// TIA Portal project "Symulacja parkingu" (V18)

(* hardware
DEVICE "S7-1200 station_1"  S7-1200 Station
   slot 0: "Rack_0"  S7-1200 Rack  Rack  V1.0
   slot 1: "PLC_1"  CPU 1214C AC/DC/Rly  6ES7 214-1BG40-0XB0  V4.6
DEVICE "HMI_1"  KTP700 Basic PN
   slot 0: "HMI_1"  KTP700 Basic PN  6AV2 123-2GB03-0AX0  17.0.0.0
   slot 1: "HMI_RT_1"  KTP700 Basic PN  6AV2 123-2GB03-0AX0  17.0.0.0
   slot 5: "HMI_1.IE_CP_1"  PROFINET Interface  17.0.0.0
      slot 1: "PROFINET Interface_1"  PROFINET Interface
         slot 1: "Port_1"  Port
*)

// ===== PLC "PLC_1"  CPU 1214C AC/DC/Rly =====

VAR_GLOBAL   // PLC tag table "Default tag table"
   "S1" AT %M0.0 : Bool;   // wjazd
   "S2" AT %M0.1 : Bool;   // wyjazd
   "S3" AT %M0.2 : Bool;   // reset
   "L1" AT %Q0.1 : Bool;   // zielone
   "L2" AT %Q0.2 : Bool;   // czerwone
   "Licznik" AT %MW10 : Word;
   "PV_Wartość_do_ustawienia" AT %MW12 : Word;
   "set wartości do ustawienia" AT %M0.3 : Bool;
   "zmienna do p_triga" AT %M0.4 : Bool;
   "S0" AT %M0.5 : Bool;   // przycisk do całkowitego wyłączenia
   "zmienna pomocnicza do przycisku od wyłączenia" AT %M0.6 : Bool;
   "całkowite wyłączenie" AT %M0.7 : Bool;
   "otwieranie szlabanu wjazd" AT %M1.0 : Bool;
   "otwieranie szlabanu wyjazd" AT %M1.1 : Bool;
   "w trakcie wyjazdu" AT %M1.2 : Bool;
   "w trakcie wjazdu" AT %M1.3 : Bool;
   "L3" AT %M1.4 : Bool;   // pomarańczowy
   "szlaban pozycja wjazd" AT %MW30 : Word;
   "szlaban podnoszenie stan wjazd" AT %M2.0 : Bool;
   "reset timera wjazd podnoszenie" AT %M2.1 : Bool;
   "szlaban opuszczania stan wjazd" AT %M2.2 : Bool;
   "reset timera wjazd opuszczanie" AT %M2.3 : Bool;
   "zmienna pomocnicza do otwierania szlabanu" AT %M2.4 : Bool;
   "szlaban pozycja wyjazd" AT %MW16 : Word;
   "szlaban podnoszenie stan wyjazd" AT %M3.0 : Bool;
   "reset timera wyjazd podnoszenie" AT %M3.1 : Bool;
   "szlaban opuszczania stan wyjazd" AT %M3.2 : Bool;
   "reset timera wyjaazd opuszcanie" AT %M3.3 : Bool;
   "zmienna pomocnicza do otwierania szlabanu 2" AT %M3.4 : Bool;
END_VAR

// folder: System blocks/Program resources

DATA_BLOCK "DB1"   // DB1
{ S7_Optimized_Access := 'TRUE' }
AUTHOR : Simatic
FAMILY : IEC
NAME : CNTR
VERSION : 1.0
// stored: InstanceOfName IEC_COUNTER
"IEC_COUNTER"
BEGIN
END_DATA_BLOCK

DATA_BLOCK "IEC_Timer_0_DB"   // DB2
{ S7_Optimized_Access := 'TRUE' }
AUTHOR : Simatic
FAMILY : IEC
NAME : IEC_TMR
VERSION : 1.0
// stored: InstanceOfName IEC_TIMER
"IEC_TIMER"
BEGIN
END_DATA_BLOCK

DATA_BLOCK "IEC_Timer_0_DB_1"   // DB3
{ S7_Optimized_Access := 'TRUE' }
AUTHOR : Simatic
FAMILY : IEC
NAME : IEC_TMR
VERSION : 1.0
// stored: InstanceOfName IEC_TIMER
"IEC_TIMER"
BEGIN
END_DATA_BLOCK

DATA_BLOCK "IEC_Timer_0_DB_2"   // DB4
{ S7_Optimized_Access := 'TRUE' }
AUTHOR : Simatic
FAMILY : IEC
NAME : IEC_TMR
VERSION : 1.0
// stored: InstanceOfName IEC_TIMER
"IEC_TIMER"
BEGIN
END_DATA_BLOCK

DATA_BLOCK "IEC_Timer_0_DB_3"   // DB5
{ S7_Optimized_Access := 'TRUE' }
AUTHOR : Simatic
FAMILY : IEC
NAME : IEC_TMR
VERSION : 1.0
// stored: InstanceOfName IEC_TIMER
"IEC_TIMER"
BEGIN
END_DATA_BLOCK

DATA_BLOCK "IEC_Timer_0_DB_4"   // DB6
{ S7_Optimized_Access := 'TRUE' }
AUTHOR : Simatic
FAMILY : IEC
NAME : IEC_TMR
VERSION : 1.0
// stored: InstanceOfName IEC_TIMER
"IEC_TIMER"
BEGIN
END_DATA_BLOCK

DATA_BLOCK "IEC_Timer_0_DB_5"   // DB7
{ S7_Optimized_Access := 'TRUE' }
AUTHOR : Simatic
FAMILY : IEC
NAME : IEC_TMR
VERSION : 1.0
// stored: InstanceOfName IEC_TIMER
"IEC_TIMER"
BEGIN
END_DATA_BLOCK

DATA_BLOCK "IEC_Timer_0_DB_6"   // DB8
{ S7_Optimized_Access := 'TRUE' }
AUTHOR : Simatic
FAMILY : IEC
NAME : IEC_TMR
VERSION : 1.0
// stored: InstanceOfName IEC_TIMER
"IEC_TIMER"
BEGIN
END_DATA_BLOCK

DATA_BLOCK "IEC_Timer_0_DB_7"   // DB9
{ S7_Optimized_Access := 'TRUE' }
AUTHOR : Simatic
FAMILY : IEC
NAME : IEC_TMR
VERSION : 1.0
// stored: InstanceOfName IEC_TIMER
"IEC_TIMER"
BEGIN
END_DATA_BLOCK

DATA_BLOCK "IEC_Timer_0_DB_8"   // DB10
{ S7_Optimized_Access := 'TRUE' }
AUTHOR : Simatic
FAMILY : IEC
NAME : IEC_TMR
VERSION : 1.0
// stored: InstanceOfName IEC_TIMER
"IEC_TIMER"
BEGIN
END_DATA_BLOCK

DATA_BLOCK "IEC_Timer_0_DB_9"   // DB11
{ S7_Optimized_Access := 'TRUE' }
AUTHOR : Simatic
FAMILY : IEC
NAME : IEC_TMR
VERSION : 1.0
// stored: InstanceOfName IEC_TIMER
"IEC_TIMER"
BEGIN
END_DATA_BLOCK

// folder: (top level)

ORGANIZATION_BLOCK "Main"   // OB1, LAD, ProgramCycle
TITLE = "Main Program Sweep (Cycle)"
{ S7_Optimized_Access := 'TRUE' }
VERSION : 0.1
   VAR_INPUT
      Initial_Call : Bool;   // Initial call of this OB
      Remanence : Bool;   // =True, if remanent data are available
   END_VAR
   VAR_TEMP   // added for the SCL form of the ladder/FBD networks
      _w1 : Bool;
   END_VAR
BEGIN

REGION Network 1
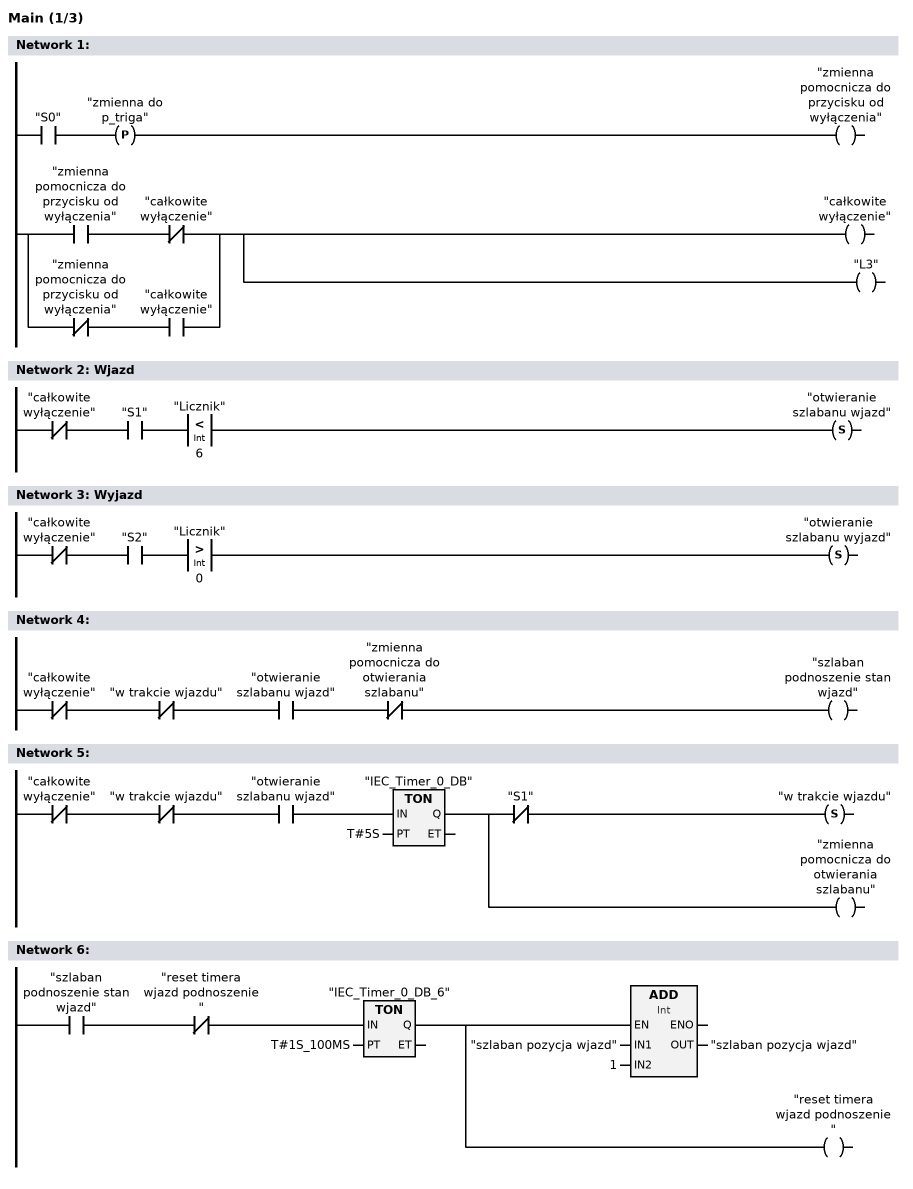
   RUNG wire#powerrail
      Contact( "S0" )
      P_Trig( "zmienna do p_triga" )
      Coil( "zmienna pomocnicza do przycisku od wyłączenia" )
   END_RUNG
   RUNG wire#powerrail
      Contact( "zmienna pomocnicza do przycisku od wyłączenia" )
      I_Contact( "całkowite wyłączenie" )
      wire#w1
      Coil( "całkowite wyłączenie" )
   END_RUNG
   RUNG wire#powerrail
      I_Contact( "zmienna pomocnicza do przycisku od wyłączenia" )
      Contact( "całkowite wyłączenie" )
   END_RUNG wire#w1
   RUNG wire#w1
      Coil( "L3" )
   END_RUNG
   // the same network as SCL:
   #_w1 := "S0" AND NOT "zmienna do p_triga";   // rising edge
   "zmienna do p_triga" := "S0";
   "zmienna pomocnicza do przycisku od wyłączenia" := #_w1;
   "całkowite wyłączenie" := ("zmienna pomocnicza do przycisku od wyłączenia" AND NOT "całkowite wyłączenie") OR (NOT "zmienna pomocnicza do przycisku od wyłączenia" AND "całkowite wyłączenie");
   "L3" := "całkowite wyłączenie";
END_REGION

REGION Network 2: Wjazd
   RUNG wire#powerrail
      I_Contact( "całkowite wyłączenie" )
      Contact( "S1" )
      { S7_Templates := "SrcType := Int" } LT_Contact(in1 := "Licznik", in2 := 6)
      S_Coil( "otwieranie szlabanu wjazd" )
   END_RUNG
   // the same network as SCL:
   IF NOT "całkowite wyłączenie" AND "S1" AND ("Licznik" < 6) THEN
       "otwieranie szlabanu wjazd" := TRUE;
   END_IF;
END_REGION

REGION Network 3: Wyjazd
   RUNG wire#powerrail
      I_Contact( "całkowite wyłączenie" )
      Contact( "S2" )
      { S7_Templates := "SrcType := Int" } GT_Contact(in1 := "Licznik", in2 := 0)
      S_Coil( "otwieranie szlabanu wyjazd" )
   END_RUNG
   // the same network as SCL:
   IF NOT "całkowite wyłączenie" AND "S2" AND ("Licznik" > 0) THEN
       "otwieranie szlabanu wyjazd" := TRUE;
   END_IF;
END_REGION

REGION Network 4
   RUNG wire#powerrail
      I_Contact( "całkowite wyłączenie" )
      I_Contact( "w trakcie wjazdu" )
      Contact( "otwieranie szlabanu wjazd" )
      I_Contact( "zmienna pomocnicza do otwierania szlabanu" )
      Coil( "szlaban podnoszenie stan wjazd" )
   END_RUNG
   // the same network as SCL:
   "szlaban podnoszenie stan wjazd" := NOT "całkowite wyłączenie" AND NOT "w trakcie wjazdu" AND "otwieranie szlabanu wjazd" AND NOT "zmienna pomocnicza do otwierania szlabanu";
END_REGION

REGION Network 5
   "IEC_Timer_0_DB".TON(IN := NOT "całkowite wyłączenie" AND NOT "w trakcie wjazdu" AND "otwieranie szlabanu wjazd",
                        PT := T#5S);
   IF "IEC_Timer_0_DB".Q AND NOT "S1" THEN "w trakcie wjazdu" := TRUE; END_IF;
   "zmienna pomocnicza do otwierania szlabanu" := "IEC_Timer_0_DB".Q;
END_REGION

REGION Network 6
   "IEC_Timer_0_DB_6".TON(IN := "szlaban podnoszenie stan wjazd" AND NOT "reset timera wjazd podnoszenie",
                          PT := T#1S_100MS);
   IF "IEC_Timer_0_DB_6".Q THEN "szlaban pozycja wjazd" := "szlaban pozycja wjazd" + 1; END_IF;
   "reset timera wjazd podnoszenie" := "IEC_Timer_0_DB_6".Q;
END_REGION

REGION Network 7
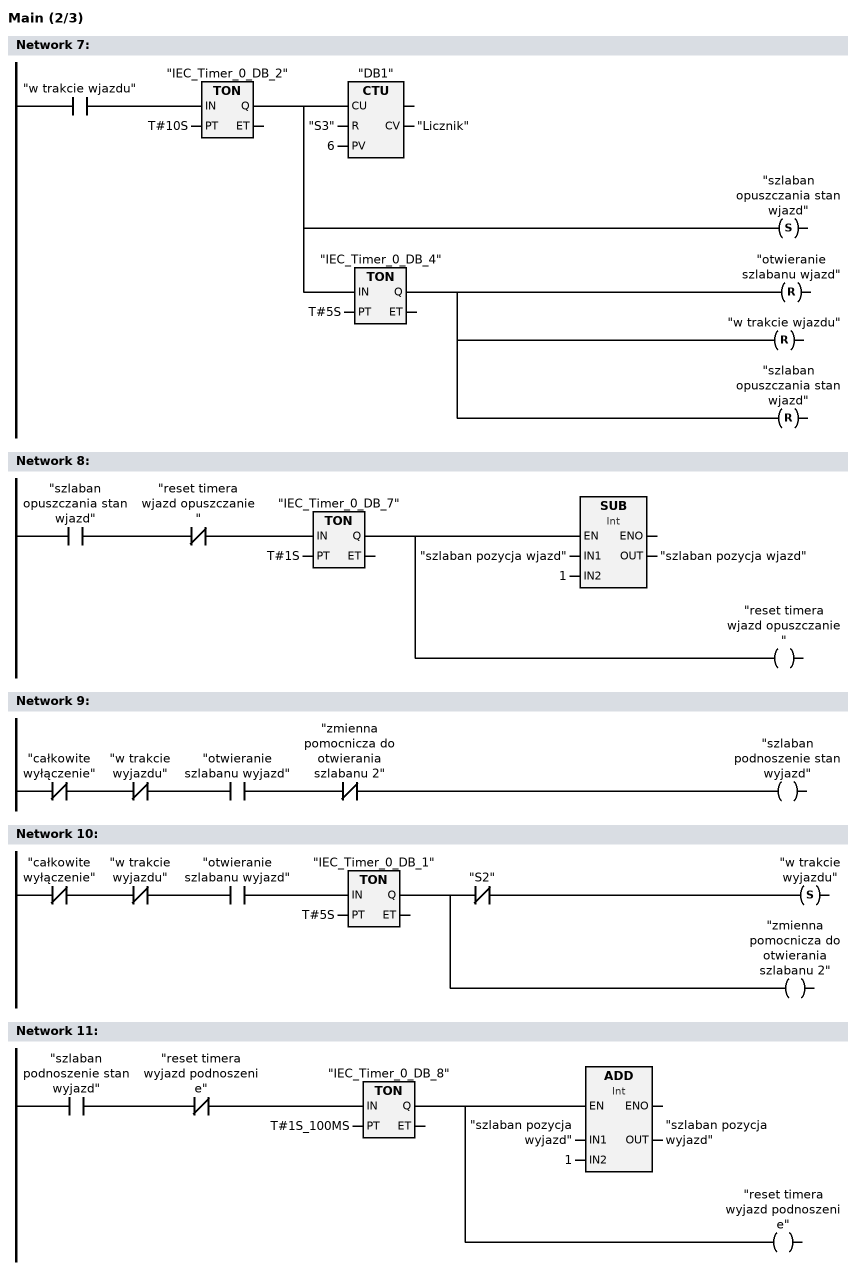
   "IEC_Timer_0_DB_2".TON(IN := "w trakcie wjazdu", PT := T#10S);
   "DB1".CTU(CU := "IEC_Timer_0_DB_2".Q, R := "S3", PV := 6, CV => "Licznik");
   IF "IEC_Timer_0_DB_2".Q THEN "szlaban opuszczania stan wjazd" := TRUE; END_IF;
   "IEC_Timer_0_DB_4".TON(IN := "IEC_Timer_0_DB_2".Q, PT := T#5S);
   IF "IEC_Timer_0_DB_4".Q THEN
       "otwieranie szlabanu wjazd" := FALSE;
       "w trakcie wjazdu" := FALSE;
       "szlaban opuszczania stan wjazd" := FALSE;
   END_IF;
END_REGION

REGION Network 8
   "IEC_Timer_0_DB_7".TON(IN := "szlaban opuszczania stan wjazd" AND NOT "reset timera wjazd opuszczanie",
                          PT := T#1S);
   IF "IEC_Timer_0_DB_7".Q THEN "szlaban pozycja wjazd" := "szlaban pozycja wjazd" - 1; END_IF;
   "reset timera wjazd opuszczanie" := "IEC_Timer_0_DB_7".Q;
END_REGION

REGION Network 9
   RUNG wire#powerrail
      I_Contact( "całkowite wyłączenie" )
      I_Contact( "w trakcie wyjazdu" )
      Contact( "otwieranie szlabanu wyjazd" )
      I_Contact( "zmienna pomocnicza do otwierania szlabanu 2" )
      Coil( "szlaban podnoszenie stan wyjazd" )
   END_RUNG
   // the same network as SCL:
   "szlaban podnoszenie stan wyjazd" := NOT "całkowite wyłączenie" AND NOT "w trakcie wyjazdu" AND "otwieranie szlabanu wyjazd" AND NOT "zmienna pomocnicza do otwierania szlabanu 2";
END_REGION

REGION Network 10
   "IEC_Timer_0_DB_1".TON(IN := NOT "całkowite wyłączenie" AND NOT "w trakcie wyjazdu" AND "otwieranie szlabanu wyjazd",
                          PT := T#5S);
   IF "IEC_Timer_0_DB_1".Q AND NOT "S2" THEN "w trakcie wyjazdu" := TRUE; END_IF;
   "zmienna pomocnicza do otwierania szlabanu 2" := "IEC_Timer_0_DB_1".Q;
END_REGION

REGION Network 11
   "IEC_Timer_0_DB_8".TON(IN := "szlaban podnoszenie stan wyjazd" AND NOT "reset timera wyjazd podnoszenie",
                          PT := T#1S_100MS);
   IF "IEC_Timer_0_DB_8".Q THEN "szlaban pozycja wyjazd" := "szlaban pozycja wyjazd" + 1; END_IF;
   "reset timera wyjazd podnoszenie" := "IEC_Timer_0_DB_8".Q;
END_REGION

REGION Network 12: wyjazd
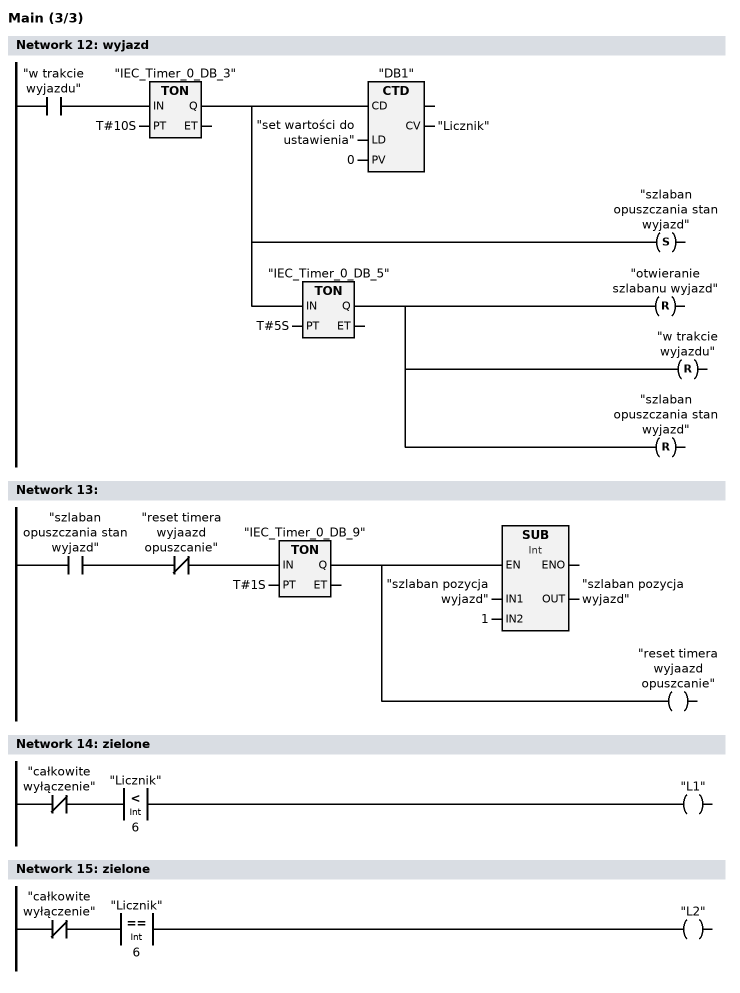
   "IEC_Timer_0_DB_3".TON(IN := "w trakcie wyjazdu", PT := T#10S);
   "DB1".CTD(CD := "IEC_Timer_0_DB_3".Q, LD := "set wartości do ustawienia", PV := 0, CV => "Licznik");
   IF "IEC_Timer_0_DB_3".Q THEN "szlaban opuszczania stan wyjazd" := TRUE; END_IF;
   "IEC_Timer_0_DB_5".TON(IN := "IEC_Timer_0_DB_3".Q, PT := T#5S);
   IF "IEC_Timer_0_DB_5".Q THEN
       "otwieranie szlabanu wyjazd" := FALSE;
       "w trakcie wyjazdu" := FALSE;
       "szlaban opuszczania stan wyjazd" := FALSE;
   END_IF;
END_REGION

REGION Network 13
   "IEC_Timer_0_DB_9".TON(IN := "szlaban opuszczania stan wyjazd" AND NOT "reset timera wyjaazd opuszcanie",
                          PT := T#1S);
   IF "IEC_Timer_0_DB_9".Q THEN "szlaban pozycja wyjazd" := "szlaban pozycja wyjazd" - 1; END_IF;
   "reset timera wyjaazd opuszcanie" := "IEC_Timer_0_DB_9".Q;
END_REGION

REGION Network 14: zielone
   RUNG wire#powerrail
      I_Contact( "całkowite wyłączenie" )
      { S7_Templates := "SrcType := Int" } LT_Contact(in1 := "Licznik", in2 := 6)
      Coil( "L1" )
   END_RUNG
   // the same network as SCL:
   "L1" := NOT "całkowite wyłączenie" AND ("Licznik" < 6);
END_REGION

REGION Network 15: zielone
   RUNG wire#powerrail
      I_Contact( "całkowite wyłączenie" )
      { S7_Templates := "SrcType := Int" } EQ_Contact(in1 := "Licznik", in2 := 6)
      Coil( "L2" )
   END_RUNG
   // the same network as SCL:
   "L2" := NOT "całkowite wyłączenie" AND ("Licznik" = 6);
END_REGION
END_ORGANIZATION_BLOCK

(* ===== HMI "HMI_RT_1" =====
system functions are stored by id; their names below are inferred from use
connection "HMI_Connection_1": ETHERNET, SMART_S7_1200_OMS

HMI tags "Default tag table"
   "Tag_ScreenNumber" : UInt, internal
   "S1" : Bool = PLC S1 AT %M0.0, 1 s
   "S2" : Bool = PLC S2 AT %M0.1, 1 s
   "Licznik" : Word = PLC Licznik AT %MW10, 1 s
   "L1" : Bool = PLC L1 AT %Q0.1, 1 s
   "L2" : Bool = PLC L2 AT %Q0.2, 1 s
   "L3" : Bool = PLC L3 AT %M1.4, 1 s
   "S3" : Bool = PLC S3 AT %M0.2, 1 s
   "S0" : Bool = PLC S0 AT %M0.5, 1 s
   "szlaban pozycja wjazd" : Word = PLC "szlaban pozycja wjazd" AT %MW30, 1 s
   "szlaban pozycja wyjazd" : Word = PLC "szlaban pozycja wyjazd" AT %MW16, 1 s

Template "Template_1" 800x480
   Button "Exit" at 714,429 size 71x50; TextOff 'Exit'; PictureOff "ExitRuntime_KTP700_Basic_PN_TR"; PictureOn "ExitRuntime_KTP700_Basic_PN_TR"
      on Release: StopRuntime(0)
   Button "Template_Button" at 614,429 size 71x50; TextOff 'Text'
   Button "Template_Button_1" at 514,429 size 71x50; TextOff 'Text'
   Button "Template_Button_2" at 414,429 size 71x50; TextOff 'Text'
   Button "Template_Button_3" at 314,429 size 71x50; TextOff 'Text'
   Button "Template_Button_4" at 214,429 size 71x50; TextOff 'Text'
   Button "Alarms" at 114,429 size 71x50; TextOff 'Alarms'; PictureOff "AlarmDisplay_KTP700_Basic_PN_TR"; PictureOn "AlarmDisplay_KTP700_Basic_PN_TR"
      on Release: function_ef3f5d25("Alarm window_Unacknowledged", -1)
   Button "Start screen" at 14,429 size 71x50; TextOff 'Start screen'; PictureOff "NavigateHome_KTP700_Basic_PN_TR"; PictureOn "NavigateHome_KTP700_Basic_PN_TR"
      on Release: ActivateScreen("Root screen", 0)
   SymbolicIOField "Symbolic_IO_Field_Screen" at 93,9 size 600x33; TextOff '0'; TextOn '1'; TextList "TextList_ScreenNames"
      ProcessValue <- "Tag_ScreenNumber"
      on Change: ActivateScreenByNumber("Tag_ScreenNumber", 0)
   DateTimeField "HmiScreenItemData" at 695,25 size 105x25
   DateTimeField "HmiScreenItemData_1" at 695,0 size 105x25
   GraphicView "Logo" at 0,0 size 91x51; Picture "Logo of HMI_1"

screen "Root screen" 800x480, template "Template_1"
   on GenerateScreen: SetTag("Tag_ScreenNumber", 1)
   TextField "HmiScreenItemData_1" at 80,225 size 640x25; Text 'Welcome to HMI_1 (KTP700 Basic+ PN)!'
   Button "HmiScreenItemData" at 36,87 size 159x47; TextOff 'Screen0'; PictureOff "Navigates to Screen0 for KTP700 Basic+ PN 17.0.0.0"; PictureOn "Navigates to Screen0 for KTP700 Basic+ PN 17.0.0.0"
      on Release: ActivateScreen("Screen0", 0)

screen "Screen0" 800x480, template "Template_1"
   on GenerateScreen: SetTag("Tag_ScreenNumber", 2)
   GraphicView "Graphic view_1" at 0,0 size 799x479
   TextField "HmiScreenItemData" at 80,225 size 640x25; Text 'Screen0'
   GraphicView "Graphic view_2" at 0,0 size 800x480; Picture "Graphic_2"
   Circle "Circle_1" at 360,295 size 48x48
      Appearance <- "L1"
   Circle "Circle_2" at 360,353 size 48x48
      Appearance <- "L2"
   Circle "Circle_3" at 360,414 size 48x48
      Appearance <- "L3"
   IOField "I/O field_1" at 338,239 size 96x32; FormatPattern 99999
      ProcessValue <- "Licznik"
   Rectangle "Rectangle_2" at 442,277 size 331x22
      VerticalMovement <- "szlaban pozycja wjazd"
   Rectangle "Rectangle_3" at 26,277 size 299x21
      VerticalMovement <- "szlaban pozycja wyjazd"
   Button "Button_1" at 564,352 size 96x32; TextOff 'Wjazd'
      Appearance <- "S1"
      on Press: SetBit("S1")
      on Release: ResetBit("S1")
   Button "Button_2" at 126,352 size 96x32; TextOff 'Wyjazd'
      Appearance <- "S2"
      on Release: ResetBit("S2")
      on Press: SetBit("S2")
   Button "Button_3" at 8,17 size 175x30; TextOff 'Reset licznika'
      Appearance <- "S3"
      on Press: SetBit("S3")
      on Release: ResetBit("S3")
   Button "Button_4" at 8,54 size 174x29; TextOff 'Wyłączenie systemu'
      Appearance <- "S0"
      on Press: SetBit("S0")
      on Release: ResetBit("S0")
*)